// TIA Portal project "Praca_Dyplomowa" (V17)

(* hardware
DEVICE "S7-1200 station_1"  S7-1200 Station
   slot 0: "Rack_0"  S7-1200 Rack  Rack  V1.0
   slot 1: "PLC_1"  CPU 1214C DC/DC/DC  6ES7 214-1AE30-0XB0  V2.2
   slot 3: "AQ 1x12BIT_1"  AQ1 signal board  6ES7 232-4HA30-0XB0  V1.0
DEVICE "HMI_2"  KTP600 Basic color PN
   slot 0: "HMI_2"  KTP600 Basic color PN  6AV6 647-0AD11-3AX0  12.0.0.0
   slot 1: "HMI_RT_2"  KTP600 Basic color PN  6AV6 647-0AD11-3AX0  12.0.0.0
   slot 5: "HMI_2.IE_CP_1"  PROFINET Interface  12.0.0.0
      slot 1: "PROFINET Interface_1"  PROFINET Interface
         slot 1: "Port_1"  Port
*)

// ===== PLC "PLC_1"  CPU 1214C DC/DC/DC =====

VAR_GLOBAL   // PLC tag table "Default tag table"
   "System_Byte" AT %MB1 : Byte;
   "FirstScan" AT %M1.0 : Bool;
   "DiagStatusUpdate" AT %M1.1 : Bool;
   "AlwaysTRUE" AT %M1.2 : Bool;
   "AlwaysFALSE" AT %M1.3 : Bool;
   "Clock_Byte" AT %MB0 : Byte;
   "Clock_10Hz" AT %M0.0 : Bool;
   "Clock_5Hz" AT %M0.1 : Bool;
   "Clock_2.5Hz" AT %M0.2 : Bool;
   "Clock_2Hz" AT %M0.3 : Bool;
   "Clock_1.25Hz" AT %M0.4 : Bool;
   "Clock_1Hz" AT %M0.5 : Bool;
   "Clock_0.625Hz" AT %M0.6 : Bool;
   "Clock_0.5Hz" AT %M0.7 : Bool;
END_VAR

DATA_BLOCK "Dane_Temperatura"   // DB1
{ S7_Optimized_Access := 'FALSE' }
VERSION : 0.1
   VAR
      DS1_DEC : Real;
      DS2_DEC : Real;
      DS3_DEC : Real;
      DS1_DECx100 : Int;
      DS2_DECx100 : Int;
      DS3_DECx100 : Int;
      Przelicznik : Real := 100.0;
      MaxDS_1 : Real;
      MinDS_1 : Real;
      MaxDS_2 : Real := 0.0;
      MinDS_2 : Real := 0.0;
      MaxDS_3 : Real := 0.0;
      MinDS_3 : Real := 0.0;
      MaxDS_1x100 : Int;
      MinDS_1x100 : Int;
      MaxDS_2x100 : Int;
      MinDS_2x100 : Int;
      MaxDS_3x100 : Int;
      MinDS_3x100 : Int;
   END_VAR
BEGIN
END_DATA_BLOCK

DATA_BLOCK "Dane Czujnik Odleglosci"   // DB2
{ S7_Optimized_Access := 'TRUE' }
VERSION : 0.1
   VAR
      Odległość : Int;
   END_VAR
BEGIN
END_DATA_BLOCK

DATA_BLOCK "MB_TCP_Data_Drugi_Serwer"   // DB4
{ S7_Optimized_Access := 'FALSE' }
VERSION : 0.1
   VAR
      IP_serwer_nr_2 : Struct
         Pierwszy_oktet : USInt := 192;
         Drugi_oktet_1 : USInt := 168;
         Trzeci_oktet_2 : USInt := 00;
         Czwarty_oktet_3 : USInt := 251;
      END_STRUCT;
      Port_Serwera_Drugiego : Word := 502;
      Serwer_Drugi : Word := 2;
      Numer_Rejestru : Word := 40001;
      Tryb_Pracy : USInt := 0;
      ILE_danych : Word := 20;
      Data_next_device : Array[1..20] of Word;
      disconnect : Bool;
      przelicznik_cisnienie : Real := 10.0;
      przelicznik_temp : Real := 100.0;
      Cisnieniex10 : Int;
      Tempx100 : Int;
      Cisnienie : Real;
      Temperatura : Real;
      Kod_Błedu : Word;
   END_VAR
BEGIN
END_DATA_BLOCK

DATA_BLOCK "MB_TCP_Data_Trzeci_Serwer"   // DB7
{ S7_Optimized_Access := 'FALSE' }
VERSION : 0.1
   VAR
      IP_serwer_nr_3 : Struct
         Pierwszy_oktet : USInt := 192;
         Drugi_oktet_1 : USInt := 168;
         Trzeci_oktet_2 : USInt := 00;
         Czwarty_oktet_3 : USInt := 252;
      END_STRUCT;
      Port_Serwera_Trzeciego : Word := 502;
      Serwer_Trzeci : Word := 3;
      Numer_Rejestru : Word := 40001;
      Tryb_Pracy : USInt := 0;
      ILE_danych : Word := 20;
      Dane_Trzeci_Serwer : Array[1..20] of Word;
      DISCONNECT : Bool;
      Kod_Błedu : Word;
      Przelicznik_100 : Real := 100.0;
      Przelicznik_1000 : Real := 1000.0;
      ax_1000 : Int;
      ay_1000 : Int;
      az_1000 : Int;
      ax : Real;
      ay : Real;
      az : Real;
      gx_100 : Int;
      gy_100 : Int;
      gz_100 : Int;
      gx : Real;
      gz : Real;
      gy : Real;
      temp_100 : Int;
      temp : Real;
   END_VAR
BEGIN
END_DATA_BLOCK

DATA_BLOCK "MB_SERWER_PLC_DANE"   // DB9
{ S7_Optimized_Access := 'FALSE' }
VERSION : 0.1
   VAR
      DISCONNECT : Bool;
      PLC_serwer_pierwszy : UInt := 5;
      IP_PORT : UInt := 502;
      New_Data_Ready : Bool;
      Data_Read : Bool;
      ERROR : Bool;
      KOD_BLEDU_SERWERA_PLC : Word;
   END_VAR
BEGIN
END_DATA_BLOCK

DATA_BLOCK "MB_TCP_Connection"   // DB10
{ S7_Optimized_Access := 'FALSE' }
VERSION : 0.1
   VAR
      MB_TCP_DISCONNECT : Bool;
      MB_TCP_ERROR : Bool;
      MB_TCP_STATUS : Word;
      MB_TCP_BUSY : Bool;
      MB_TCP_DONE : Bool;
      Connection_Lost : Bool;
   END_VAR
BEGIN
END_DATA_BLOCK

DATA_BLOCK "MB_TCP_Data"   // DB11
{ S7_Optimized_Access := 'FALSE' }
VERSION : 0.1
   VAR
      IP_serwer_nr_1 : Struct
         Pierwszy_oktet : USInt := 192;
         Drugi_oktet_1 : USInt := 168;
         Trzeci_oktet_2 : USInt := 00;
         Czwarty_oktet_3 : USInt := 253;
      END_STRUCT;
      Port_Serwera_Pierwszego : Word := 502;
      Serwer_Pierwszy : Word := 1;
      Numer_Rejestru : Word := 40001;
      Tryb_Pracy : USInt := 0;
      ILE_danych : Word := 26;
      Dane_serwer_pierwszy : Array[1..26] of Word;
   END_VAR
BEGIN
END_DATA_BLOCK

DATA_BLOCK "Zmienne_cyclic_interrupt"   // DB12
{ S7_Optimized_Access := 'TRUE' }
VERSION : 0.1
   VAR RETAIN
      IN : Bool;
      PIN : Bool;
      OUT : Bool;
      POUT : Bool;
      Czas : Time := T#250ms;
   END_VAR
BEGIN
END_DATA_BLOCK

FUNCTION "VL53L1" : Void   // FC1, LAD
{ S7_Optimized_Access := 'TRUE' }
VERSION : 0.1
BEGIN

REGION Network 1
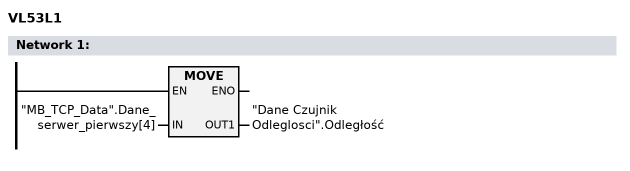
   RUNG wire#powerrail
      { S7_GenerateENO := "TRUE" } Move(in := "MB_TCP_Data".Dane_serwer_pierwszy[4], out1 => "Dane Czujnik Odleglosci".Odległość)
   END_RUNG
   // the same network as SCL:
   "Dane Czujnik Odleglosci".Odległość := "MB_TCP_Data".Dane_serwer_pierwszy[4];
END_REGION
END_FUNCTION

FUNCTION "STATUS_INFO" : Void   // FC2, SCL
{ S7_Optimized_Access := 'TRUE' }
VERSION : 0.1
   VAR_TEMP
      i : Int;
      "a" : Int;
      "b" : Int;
   END_VAR
BEGIN
   IF WORD_TO_INT("MB_TCP_Connection".MB_TCP_STATUS) <> 0 THEN
       "MB_TCP_Connection".Connection_Lost := TRUE;
       FOR #i := 1 TO WORD_TO_INT("MB_TCP_Data".ILE_danych) DO
           "MB_TCP_Data".Dane_serwer_pierwszy[#i] := 0;
       END_FOR;
   ELSE
       "MB_TCP_Connection".Connection_Lost := FALSE;
   END_IF;

   IF WORD_TO_INT("MB_TCP_Data_Drugi_Serwer".Kod_Błedu) <> 0 THEN

       FOR #a := 1 TO WORD_TO_INT("MB_TCP_Data_Trzeci_Serwer".ILE_danych) DO
           "MB_TCP_Data_Drugi_Serwer".Data_next_device[#a] := 0;
       END_FOR;

   END_IF;


   IF WORD_TO_INT("MB_TCP_Data_Trzeci_Serwer".Kod_Błedu) <> 0 THEN

       FOR #b := 1 TO WORD_TO_INT("MB_TCP_Data_Trzeci_Serwer".ILE_danych) DO
           "MB_TCP_Data_Trzeci_Serwer".Dane_Trzeci_Serwer[#b] := 0;
       END_FOR;

   END_IF;
END_FUNCTION

FUNCTION "BMP280" : Void   // FC3, LAD
{ S7_Optimized_Access := 'TRUE' }
VERSION : 0.1
BEGIN

REGION Network 1
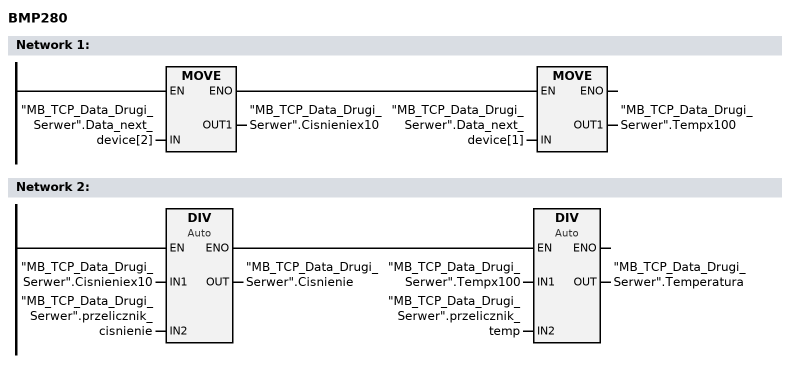
   RUNG wire#powerrail
      { S7_GenerateENO := "TRUE" } Move(in := "MB_TCP_Data_Drugi_Serwer".Data_next_device[2], out1 => "MB_TCP_Data_Drugi_Serwer".Cisnieniex10)
      { S7_GenerateENO := "TRUE" } Move(in := "MB_TCP_Data_Drugi_Serwer".Data_next_device[1], out1 => "MB_TCP_Data_Drugi_Serwer".Tempx100)
   END_RUNG
   // the same network as SCL:
   // ENO of a box is taken as its EN; it also drops when the box reports an error
   "MB_TCP_Data_Drugi_Serwer".Cisnieniex10 := "MB_TCP_Data_Drugi_Serwer".Data_next_device[2];
   "MB_TCP_Data_Drugi_Serwer".Tempx100 := "MB_TCP_Data_Drugi_Serwer".Data_next_device[1];
END_REGION

REGION Network 2
   RUNG wire#powerrail
      { S7_GenerateENO := "TRUE" } Div(in1 := "MB_TCP_Data_Drugi_Serwer".Cisnieniex10, in2 := "MB_TCP_Data_Drugi_Serwer".przelicznik_cisnienie, out => "MB_TCP_Data_Drugi_Serwer".Cisnienie)
      { S7_GenerateENO := "TRUE" } Div(in1 := "MB_TCP_Data_Drugi_Serwer".Tempx100, in2 := "MB_TCP_Data_Drugi_Serwer".przelicznik_temp, out => "MB_TCP_Data_Drugi_Serwer".Temperatura)
   END_RUNG
   // the same network as SCL:
   // ENO of a box is taken as its EN; it also drops when the box reports an error
   "MB_TCP_Data_Drugi_Serwer".Cisnienie := "MB_TCP_Data_Drugi_Serwer".Cisnieniex10 / "MB_TCP_Data_Drugi_Serwer".przelicznik_cisnienie;
   "MB_TCP_Data_Drugi_Serwer".Temperatura := "MB_TCP_Data_Drugi_Serwer".Tempx100 / "MB_TCP_Data_Drugi_Serwer".przelicznik_temp;
END_REGION
END_FUNCTION

FUNCTION "GY521" : Void   // FC4, LAD
{ S7_Optimized_Access := 'TRUE' }
VERSION : 0.1
BEGIN

REGION Network 1
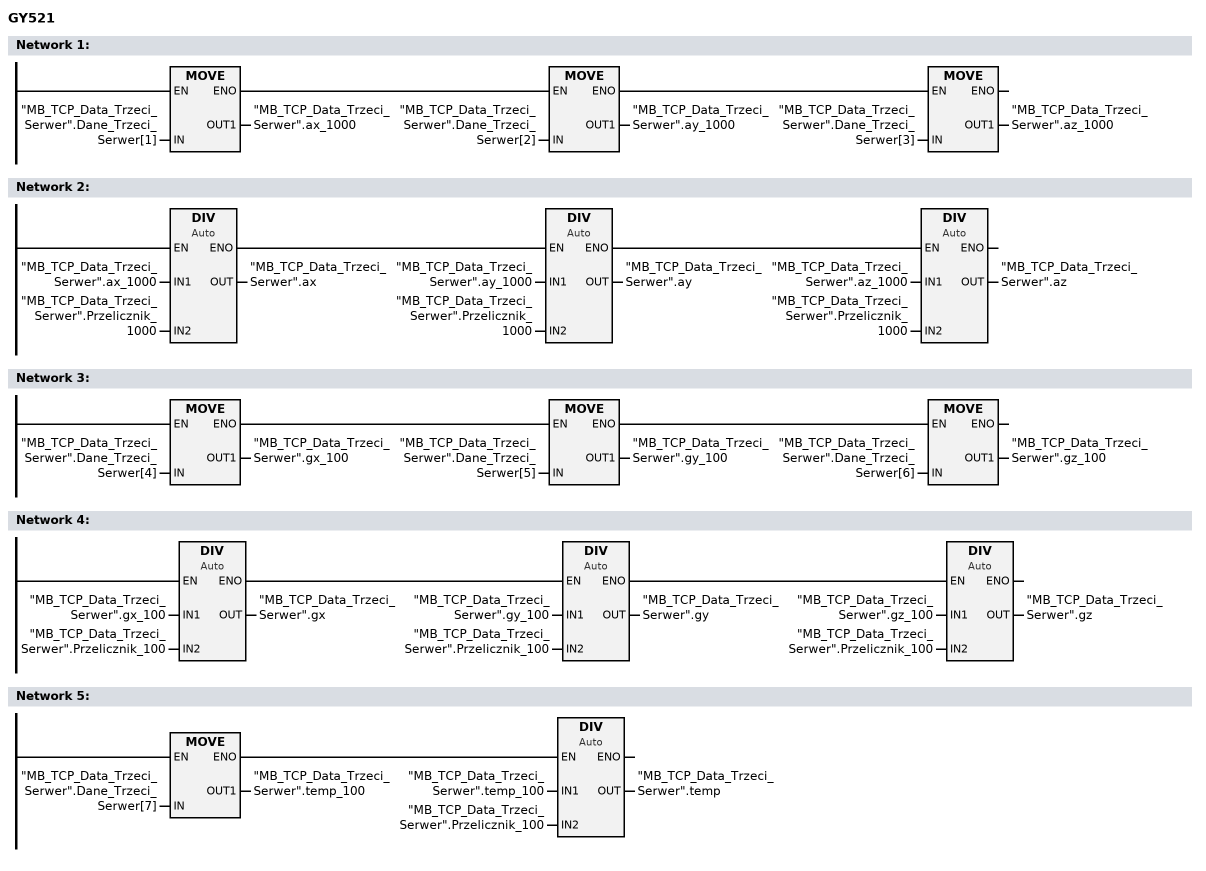
   RUNG wire#powerrail
      { S7_GenerateENO := "TRUE" } Move(in := "MB_TCP_Data_Trzeci_Serwer".Dane_Trzeci_Serwer[1], out1 => "MB_TCP_Data_Trzeci_Serwer".ax_1000)
      { S7_GenerateENO := "TRUE" } Move(in := "MB_TCP_Data_Trzeci_Serwer".Dane_Trzeci_Serwer[2], out1 => "MB_TCP_Data_Trzeci_Serwer".ay_1000)
      { S7_GenerateENO := "TRUE" } Move(in := "MB_TCP_Data_Trzeci_Serwer".Dane_Trzeci_Serwer[3], out1 => "MB_TCP_Data_Trzeci_Serwer".az_1000)
   END_RUNG
   // the same network as SCL:
   // ENO of a box is taken as its EN; it also drops when the box reports an error
   "MB_TCP_Data_Trzeci_Serwer".ax_1000 := "MB_TCP_Data_Trzeci_Serwer".Dane_Trzeci_Serwer[1];
   "MB_TCP_Data_Trzeci_Serwer".ay_1000 := "MB_TCP_Data_Trzeci_Serwer".Dane_Trzeci_Serwer[2];
   "MB_TCP_Data_Trzeci_Serwer".az_1000 := "MB_TCP_Data_Trzeci_Serwer".Dane_Trzeci_Serwer[3];
END_REGION

REGION Network 2
   RUNG wire#powerrail
      { S7_GenerateENO := "TRUE" } Div(in1 := "MB_TCP_Data_Trzeci_Serwer".ax_1000, in2 := "MB_TCP_Data_Trzeci_Serwer".Przelicznik_1000, out => "MB_TCP_Data_Trzeci_Serwer".ax)
      { S7_GenerateENO := "TRUE" } Div(in1 := "MB_TCP_Data_Trzeci_Serwer".ay_1000, in2 := "MB_TCP_Data_Trzeci_Serwer".Przelicznik_1000, out => "MB_TCP_Data_Trzeci_Serwer".ay)
      { S7_GenerateENO := "TRUE" } Div(in1 := "MB_TCP_Data_Trzeci_Serwer".az_1000, in2 := "MB_TCP_Data_Trzeci_Serwer".Przelicznik_1000, out => "MB_TCP_Data_Trzeci_Serwer".az)
   END_RUNG
   // the same network as SCL:
   // ENO of a box is taken as its EN; it also drops when the box reports an error
   "MB_TCP_Data_Trzeci_Serwer".ax := "MB_TCP_Data_Trzeci_Serwer".ax_1000 / "MB_TCP_Data_Trzeci_Serwer".Przelicznik_1000;
   "MB_TCP_Data_Trzeci_Serwer".ay := "MB_TCP_Data_Trzeci_Serwer".ay_1000 / "MB_TCP_Data_Trzeci_Serwer".Przelicznik_1000;
   "MB_TCP_Data_Trzeci_Serwer".az := "MB_TCP_Data_Trzeci_Serwer".az_1000 / "MB_TCP_Data_Trzeci_Serwer".Przelicznik_1000;
END_REGION

REGION Network 3
   RUNG wire#powerrail
      { S7_GenerateENO := "TRUE" } Move(in := "MB_TCP_Data_Trzeci_Serwer".Dane_Trzeci_Serwer[4], out1 => "MB_TCP_Data_Trzeci_Serwer".gx_100)
      { S7_GenerateENO := "TRUE" } Move(in := "MB_TCP_Data_Trzeci_Serwer".Dane_Trzeci_Serwer[5], out1 => "MB_TCP_Data_Trzeci_Serwer".gy_100)
      { S7_GenerateENO := "TRUE" } Move(in := "MB_TCP_Data_Trzeci_Serwer".Dane_Trzeci_Serwer[6], out1 => "MB_TCP_Data_Trzeci_Serwer".gz_100)
   END_RUNG
   // the same network as SCL:
   // ENO of a box is taken as its EN; it also drops when the box reports an error
   "MB_TCP_Data_Trzeci_Serwer".gx_100 := "MB_TCP_Data_Trzeci_Serwer".Dane_Trzeci_Serwer[4];
   "MB_TCP_Data_Trzeci_Serwer".gy_100 := "MB_TCP_Data_Trzeci_Serwer".Dane_Trzeci_Serwer[5];
   "MB_TCP_Data_Trzeci_Serwer".gz_100 := "MB_TCP_Data_Trzeci_Serwer".Dane_Trzeci_Serwer[6];
END_REGION

REGION Network 4
   RUNG wire#powerrail
      { S7_GenerateENO := "TRUE" } Div(in1 := "MB_TCP_Data_Trzeci_Serwer".gx_100, in2 := "MB_TCP_Data_Trzeci_Serwer".Przelicznik_100, out => "MB_TCP_Data_Trzeci_Serwer".gx)
      { S7_GenerateENO := "TRUE" } Div(in1 := "MB_TCP_Data_Trzeci_Serwer".gy_100, in2 := "MB_TCP_Data_Trzeci_Serwer".Przelicznik_100, out => "MB_TCP_Data_Trzeci_Serwer".gy)
      { S7_GenerateENO := "TRUE" } Div(in1 := "MB_TCP_Data_Trzeci_Serwer".gz_100, in2 := "MB_TCP_Data_Trzeci_Serwer".Przelicznik_100, out => "MB_TCP_Data_Trzeci_Serwer".gz)
   END_RUNG
   // the same network as SCL:
   // ENO of a box is taken as its EN; it also drops when the box reports an error
   "MB_TCP_Data_Trzeci_Serwer".gx := "MB_TCP_Data_Trzeci_Serwer".gx_100 / "MB_TCP_Data_Trzeci_Serwer".Przelicznik_100;
   "MB_TCP_Data_Trzeci_Serwer".gy := "MB_TCP_Data_Trzeci_Serwer".gy_100 / "MB_TCP_Data_Trzeci_Serwer".Przelicznik_100;
   "MB_TCP_Data_Trzeci_Serwer".gz := "MB_TCP_Data_Trzeci_Serwer".gz_100 / "MB_TCP_Data_Trzeci_Serwer".Przelicznik_100;
END_REGION

REGION Network 5
   RUNG wire#powerrail
      { S7_GenerateENO := "TRUE" } Move(in := "MB_TCP_Data_Trzeci_Serwer".Dane_Trzeci_Serwer[7], out1 => "MB_TCP_Data_Trzeci_Serwer".temp_100)
      { S7_GenerateENO := "TRUE" } Div(in1 := "MB_TCP_Data_Trzeci_Serwer".temp_100, in2 := "MB_TCP_Data_Trzeci_Serwer".Przelicznik_100, out => "MB_TCP_Data_Trzeci_Serwer".temp)
   END_RUNG
   // the same network as SCL:
   // ENO of a box is taken as its EN; it also drops when the box reports an error
   "MB_TCP_Data_Trzeci_Serwer".temp_100 := "MB_TCP_Data_Trzeci_Serwer".Dane_Trzeci_Serwer[7];
   "MB_TCP_Data_Trzeci_Serwer".temp := "MB_TCP_Data_Trzeci_Serwer".temp_100 / "MB_TCP_Data_Trzeci_Serwer".Przelicznik_100;
END_REGION
END_FUNCTION

FUNCTION "MB_Serwer_PLC" : Void   // FC5, LAD
{ S7_Optimized_Access := 'FALSE' }
VERSION : 0.1
BEGIN

REGION Network 1
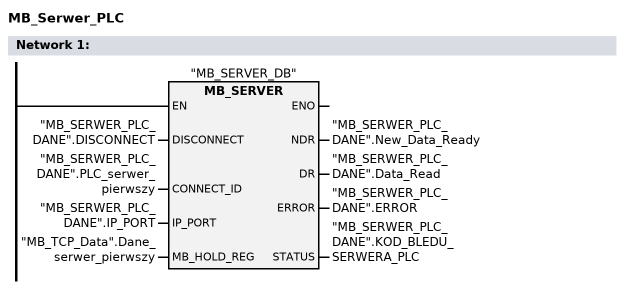
   "MB_SERVER_DB"(DISCONNECT := "MB_SERWER_PLC_DANE".DISCONNECT,   // MB_SERVER
                  CONNECT_ID := "MB_SERWER_PLC_DANE".PLC_serwer_pierwszy,
                  IP_PORT := "MB_SERWER_PLC_DANE".IP_PORT,
                  MB_HOLD_REG := "MB_TCP_Data".Dane_serwer_pierwszy,
                  NDR => "MB_SERWER_PLC_DANE".New_Data_Ready,
                  DR => "MB_SERWER_PLC_DANE".Data_Read,
                  ERROR => "MB_SERWER_PLC_DANE".ERROR,
                  STATUS => "MB_SERWER_PLC_DANE".KOD_BLEDU_SERWERA_PLC);
END_REGION
END_FUNCTION

FUNCTION "FC_BMTCP_Client" : Void   // FC10, LAD
{ S7_Optimized_Access := 'FALSE' }
VERSION : 0.1
BEGIN

REGION Network 1
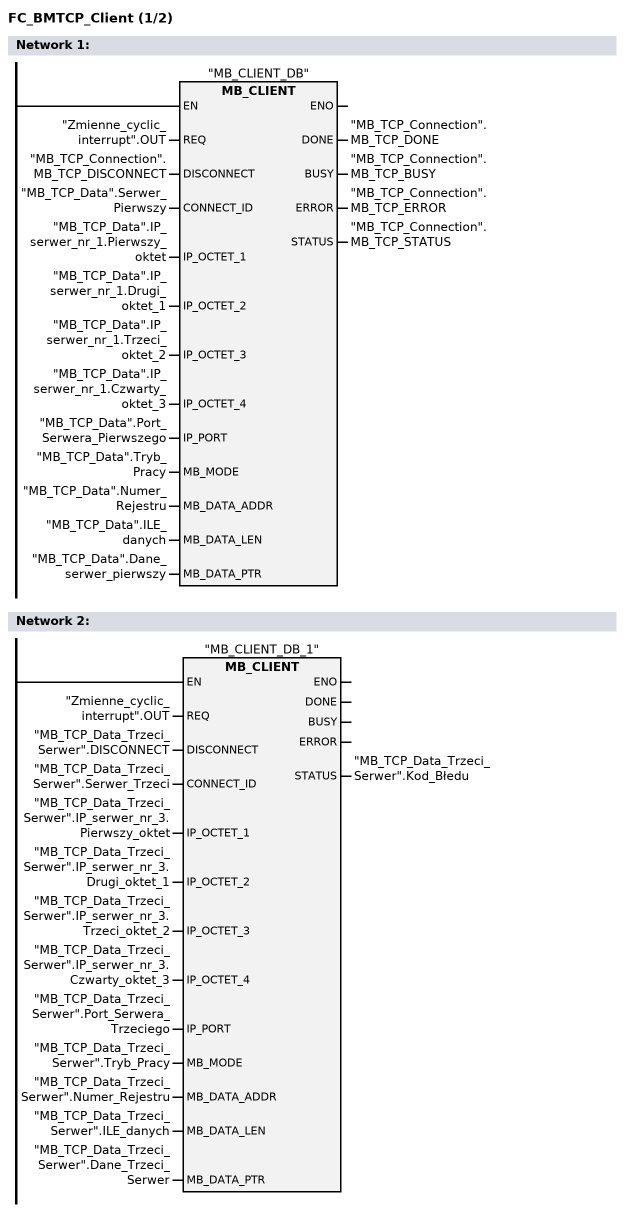
   "MB_CLIENT_DB"(REQ := "Zmienne_cyclic_interrupt".OUT,   // MB_CLIENT
                  DISCONNECT := "MB_TCP_Connection".MB_TCP_DISCONNECT,
                  CONNECT_ID := "MB_TCP_Data".Serwer_Pierwszy,
                  IP_OCTET_1 := "MB_TCP_Data".IP_serwer_nr_1.Pierwszy_oktet,
                  IP_OCTET_2 := "MB_TCP_Data".IP_serwer_nr_1.Drugi_oktet_1,
                  IP_OCTET_3 := "MB_TCP_Data".IP_serwer_nr_1.Trzeci_oktet_2,
                  IP_OCTET_4 := "MB_TCP_Data".IP_serwer_nr_1.Czwarty_oktet_3,
                  IP_PORT := "MB_TCP_Data".Port_Serwera_Pierwszego,
                  MB_MODE := "MB_TCP_Data".Tryb_Pracy,
                  MB_DATA_ADDR := "MB_TCP_Data".Numer_Rejestru,
                  MB_DATA_LEN := "MB_TCP_Data".ILE_danych,
                  MB_DATA_PTR := "MB_TCP_Data".Dane_serwer_pierwszy,
                  DONE => "MB_TCP_Connection".MB_TCP_DONE,
                  BUSY => "MB_TCP_Connection".MB_TCP_BUSY,
                  ERROR => "MB_TCP_Connection".MB_TCP_ERROR,
                  STATUS => "MB_TCP_Connection".MB_TCP_STATUS);
END_REGION

REGION Network 2
   "MB_CLIENT_DB_1"(REQ := "Zmienne_cyclic_interrupt".OUT,   // MB_CLIENT
                    DISCONNECT := "MB_TCP_Data_Trzeci_Serwer".DISCONNECT,
                    CONNECT_ID := "MB_TCP_Data_Trzeci_Serwer".Serwer_Trzeci,
                    IP_OCTET_1 := "MB_TCP_Data_Trzeci_Serwer".IP_serwer_nr_3.Pierwszy_oktet,
                    IP_OCTET_2 := "MB_TCP_Data_Trzeci_Serwer".IP_serwer_nr_3.Drugi_oktet_1,
                    IP_OCTET_3 := "MB_TCP_Data_Trzeci_Serwer".IP_serwer_nr_3.Trzeci_oktet_2,
                    IP_OCTET_4 := "MB_TCP_Data_Trzeci_Serwer".IP_serwer_nr_3.Czwarty_oktet_3,
                    IP_PORT := "MB_TCP_Data_Trzeci_Serwer".Port_Serwera_Trzeciego,
                    MB_MODE := "MB_TCP_Data_Trzeci_Serwer".Tryb_Pracy,
                    MB_DATA_ADDR := "MB_TCP_Data_Trzeci_Serwer".Numer_Rejestru,
                    MB_DATA_LEN := "MB_TCP_Data_Trzeci_Serwer".ILE_danych,
                    MB_DATA_PTR := "MB_TCP_Data_Trzeci_Serwer".Dane_Trzeci_Serwer,
                    STATUS => "MB_TCP_Data_Trzeci_Serwer".Kod_Błedu);
END_REGION

REGION Network 3
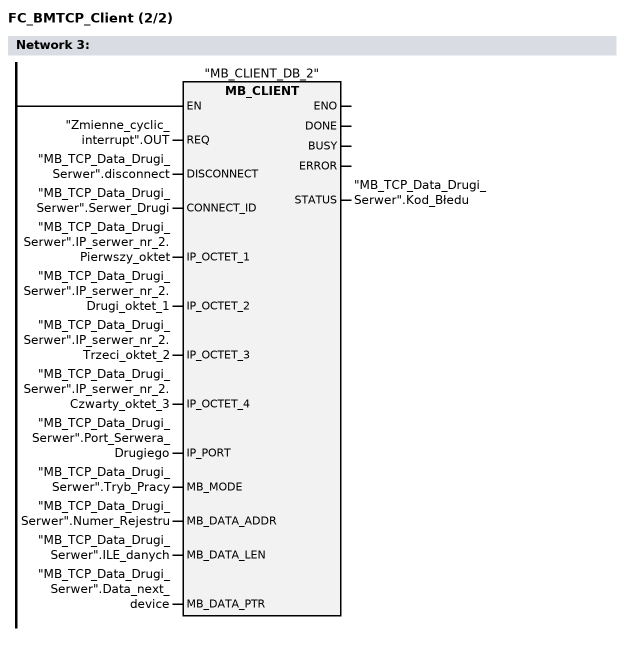
   "MB_CLIENT_DB_2"(REQ := "Zmienne_cyclic_interrupt".OUT,   // MB_CLIENT
                    DISCONNECT := "MB_TCP_Data_Drugi_Serwer".disconnect,
                    CONNECT_ID := "MB_TCP_Data_Drugi_Serwer".Serwer_Drugi,
                    IP_OCTET_1 := "MB_TCP_Data_Drugi_Serwer".IP_serwer_nr_2.Pierwszy_oktet,
                    IP_OCTET_2 := "MB_TCP_Data_Drugi_Serwer".IP_serwer_nr_2.Drugi_oktet_1,
                    IP_OCTET_3 := "MB_TCP_Data_Drugi_Serwer".IP_serwer_nr_2.Trzeci_oktet_2,
                    IP_OCTET_4 := "MB_TCP_Data_Drugi_Serwer".IP_serwer_nr_2.Czwarty_oktet_3,
                    IP_PORT := "MB_TCP_Data_Drugi_Serwer".Port_Serwera_Drugiego,
                    MB_MODE := "MB_TCP_Data_Drugi_Serwer".Tryb_Pracy,
                    MB_DATA_ADDR := "MB_TCP_Data_Drugi_Serwer".Numer_Rejestru,
                    MB_DATA_LEN := "MB_TCP_Data_Drugi_Serwer".ILE_danych,
                    MB_DATA_PTR := "MB_TCP_Data_Drugi_Serwer".Data_next_device,
                    STATUS => "MB_TCP_Data_Drugi_Serwer".Kod_Błedu);
END_REGION
END_FUNCTION

FUNCTION "TEMP_HEX_AND_REAL" : Void   // FC11, LAD
{ S7_Optimized_Access := 'FALSE' }
VERSION : 0.1
BEGIN

REGION Network 1
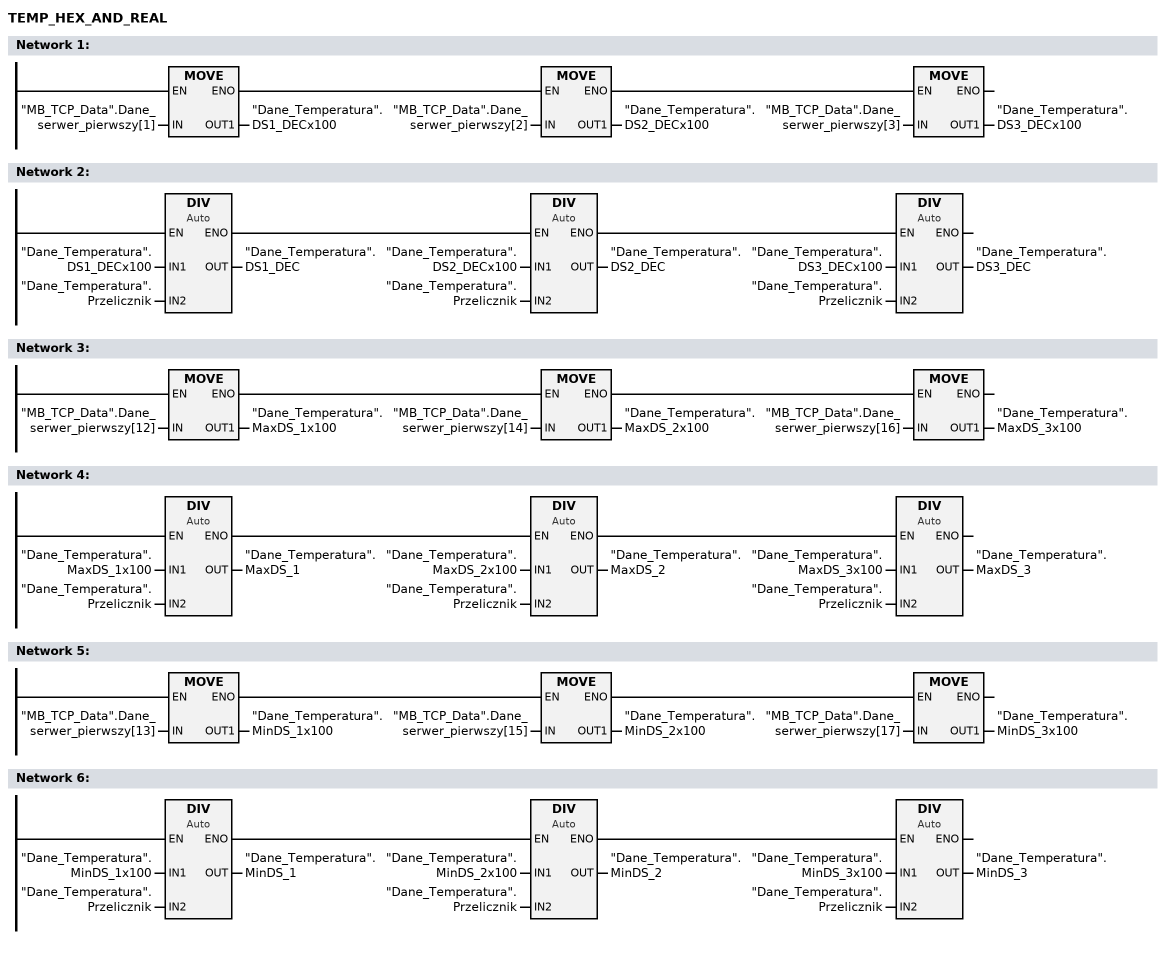
   RUNG wire#powerrail
      { S7_GenerateENO := "TRUE" } Move(in := "MB_TCP_Data".Dane_serwer_pierwszy[1], out1 => "Dane_Temperatura".DS1_DECx100)
      { S7_GenerateENO := "TRUE" } Move(in := "MB_TCP_Data".Dane_serwer_pierwszy[2], out1 => "Dane_Temperatura".DS2_DECx100)
      { S7_GenerateENO := "TRUE" } Move(in := "MB_TCP_Data".Dane_serwer_pierwszy[3], out1 => "Dane_Temperatura".DS3_DECx100)
   END_RUNG
   // the same network as SCL:
   // ENO of a box is taken as its EN; it also drops when the box reports an error
   "Dane_Temperatura".DS1_DECx100 := "MB_TCP_Data".Dane_serwer_pierwszy[1];
   "Dane_Temperatura".DS2_DECx100 := "MB_TCP_Data".Dane_serwer_pierwszy[2];
   "Dane_Temperatura".DS3_DECx100 := "MB_TCP_Data".Dane_serwer_pierwszy[3];
END_REGION

REGION Network 2
   RUNG wire#powerrail
      { S7_GenerateENO := "TRUE" } Div(in1 := "Dane_Temperatura".DS1_DECx100, in2 := "Dane_Temperatura".Przelicznik, out => "Dane_Temperatura".DS1_DEC)
      { S7_GenerateENO := "TRUE" } Div(in1 := "Dane_Temperatura".DS2_DECx100, in2 := "Dane_Temperatura".Przelicznik, out => "Dane_Temperatura".DS2_DEC)
      { S7_GenerateENO := "TRUE" } Div(in1 := "Dane_Temperatura".DS3_DECx100, in2 := "Dane_Temperatura".Przelicznik, out => "Dane_Temperatura".DS3_DEC)
   END_RUNG
   // the same network as SCL:
   // ENO of a box is taken as its EN; it also drops when the box reports an error
   "Dane_Temperatura".DS1_DEC := "Dane_Temperatura".DS1_DECx100 / "Dane_Temperatura".Przelicznik;
   "Dane_Temperatura".DS2_DEC := "Dane_Temperatura".DS2_DECx100 / "Dane_Temperatura".Przelicznik;
   "Dane_Temperatura".DS3_DEC := "Dane_Temperatura".DS3_DECx100 / "Dane_Temperatura".Przelicznik;
END_REGION

REGION Network 3
   RUNG wire#powerrail
      { S7_GenerateENO := "TRUE" } Move(in := "MB_TCP_Data".Dane_serwer_pierwszy[12], out1 => "Dane_Temperatura".MaxDS_1x100)
      { S7_GenerateENO := "TRUE" } Move(in := "MB_TCP_Data".Dane_serwer_pierwszy[14], out1 => "Dane_Temperatura".MaxDS_2x100)
      { S7_GenerateENO := "TRUE" } Move(in := "MB_TCP_Data".Dane_serwer_pierwszy[16], out1 => "Dane_Temperatura".MaxDS_3x100)
   END_RUNG
   // the same network as SCL:
   // ENO of a box is taken as its EN; it also drops when the box reports an error
   "Dane_Temperatura".MaxDS_1x100 := "MB_TCP_Data".Dane_serwer_pierwszy[12];
   "Dane_Temperatura".MaxDS_2x100 := "MB_TCP_Data".Dane_serwer_pierwszy[14];
   "Dane_Temperatura".MaxDS_3x100 := "MB_TCP_Data".Dane_serwer_pierwszy[16];
END_REGION

REGION Network 4
   RUNG wire#powerrail
      { S7_GenerateENO := "TRUE" } Div(in1 := "Dane_Temperatura".MaxDS_1x100, in2 := "Dane_Temperatura".Przelicznik, out => "Dane_Temperatura".MaxDS_1)
      { S7_GenerateENO := "TRUE" } Div(in1 := "Dane_Temperatura".MaxDS_2x100, in2 := "Dane_Temperatura".Przelicznik, out => "Dane_Temperatura".MaxDS_2)
      { S7_GenerateENO := "TRUE" } Div(in1 := "Dane_Temperatura".MaxDS_3x100, in2 := "Dane_Temperatura".Przelicznik, out => "Dane_Temperatura".MaxDS_3)
   END_RUNG
   // the same network as SCL:
   // ENO of a box is taken as its EN; it also drops when the box reports an error
   "Dane_Temperatura".MaxDS_1 := "Dane_Temperatura".MaxDS_1x100 / "Dane_Temperatura".Przelicznik;
   "Dane_Temperatura".MaxDS_2 := "Dane_Temperatura".MaxDS_2x100 / "Dane_Temperatura".Przelicznik;
   "Dane_Temperatura".MaxDS_3 := "Dane_Temperatura".MaxDS_3x100 / "Dane_Temperatura".Przelicznik;
END_REGION

REGION Network 5
   RUNG wire#powerrail
      { S7_GenerateENO := "TRUE" } Move(in := "MB_TCP_Data".Dane_serwer_pierwszy[13], out1 => "Dane_Temperatura".MinDS_1x100)
      { S7_GenerateENO := "TRUE" } Move(in := "MB_TCP_Data".Dane_serwer_pierwszy[15], out1 => "Dane_Temperatura".MinDS_2x100)
      { S7_GenerateENO := "TRUE" } Move(in := "MB_TCP_Data".Dane_serwer_pierwszy[17], out1 => "Dane_Temperatura".MinDS_3x100)
   END_RUNG
   // the same network as SCL:
   // ENO of a box is taken as its EN; it also drops when the box reports an error
   "Dane_Temperatura".MinDS_1x100 := "MB_TCP_Data".Dane_serwer_pierwszy[13];
   "Dane_Temperatura".MinDS_2x100 := "MB_TCP_Data".Dane_serwer_pierwszy[15];
   "Dane_Temperatura".MinDS_3x100 := "MB_TCP_Data".Dane_serwer_pierwszy[17];
END_REGION

REGION Network 6
   RUNG wire#powerrail
      { S7_GenerateENO := "TRUE" } Div(in1 := "Dane_Temperatura".MinDS_1x100, in2 := "Dane_Temperatura".Przelicznik, out => "Dane_Temperatura".MinDS_1)
      { S7_GenerateENO := "TRUE" } Div(in1 := "Dane_Temperatura".MinDS_2x100, in2 := "Dane_Temperatura".Przelicznik, out => "Dane_Temperatura".MinDS_2)
      { S7_GenerateENO := "TRUE" } Div(in1 := "Dane_Temperatura".MinDS_3x100, in2 := "Dane_Temperatura".Przelicznik, out => "Dane_Temperatura".MinDS_3)
   END_RUNG
   // the same network as SCL:
   // ENO of a box is taken as its EN; it also drops when the box reports an error
   "Dane_Temperatura".MinDS_1 := "Dane_Temperatura".MinDS_1x100 / "Dane_Temperatura".Przelicznik;
   "Dane_Temperatura".MinDS_2 := "Dane_Temperatura".MinDS_2x100 / "Dane_Temperatura".Przelicznik;
   "Dane_Temperatura".MinDS_3 := "Dane_Temperatura".MinDS_3x100 / "Dane_Temperatura".Przelicznik;
END_REGION
END_FUNCTION

ORGANIZATION_BLOCK "Main"   // OB1, LAD, ProgramCycle
TITLE = "Main Program Sweep (Cycle)"
{ S7_Optimized_Access := 'TRUE' }
VERSION : 0.1
   VAR_TEMP   // added for the SCL form of the ladder/FBD networks
      _w1 : Bool;
      _w2 : Bool;
      _w3 : Bool;
      _w4 : Bool;
      _w5 : Bool;
   END_VAR
BEGIN

REGION Network 1
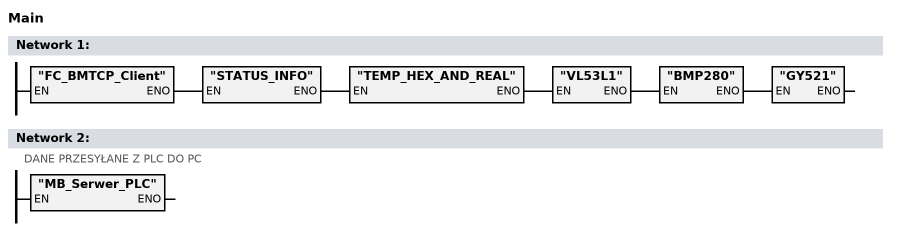
   RUNG wire#powerrail
      "FC_BMTCP_Client"()
      "STATUS_INFO"()
      "TEMP_HEX_AND_REAL"()
      "VL53L1"()
      "BMP280"()
      "GY521"()
   END_RUNG
   // the same network as SCL:
   "FC_BMTCP_Client"(ENO => #_w1);
   "STATUS_INFO"(EN := #_w1, ENO => #_w2);
   "TEMP_HEX_AND_REAL"(EN := #_w2, ENO => #_w3);
   "VL53L1"(EN := #_w3, ENO => #_w4);
   "BMP280"(EN := #_w4, ENO => #_w5);
   IF #_w5 THEN "GY521"(); END_IF;
END_REGION

REGION Network 2
   // DANE PRZESYŁANE Z PLC DO PC
   RUNG wire#powerrail
      "MB_Serwer_PLC"()
   END_RUNG
   // the same network as SCL:
   "MB_Serwer_PLC"();
END_REGION
END_ORGANIZATION_BLOCK

ORGANIZATION_BLOCK "Cyclic interrupt"   // OB30, SCL, CyclicInterrupt
{ S7_Optimized_Access := 'TRUE' }
VERSION : 0.1
BEGIN
   "Zmienne_cyclic_interrupt".OUT := NOT "Zmienne_cyclic_interrupt".OUT;
END_ORGANIZATION_BLOCK

(* ===== HMI "HMI_RT_2" =====
system functions are stored by id; their names below are inferred from use
connection "HMI_Connection_2": ETHERNET, SMART_S7_1200_OMS

HMI tags "Default tag table"
   "Dane_Temperatura_DS1_DEC" : Real = PLC Dane_Temperatura.DS1_DEC AT %DB1.DBD0, 100 ms
   "Dane_Temperatura_DS2_DEC" : Real = PLC Dane_Temperatura.DS2_DEC AT %DB1.DBD4, 100 ms
   "Dane_Temperatura_DS3_DEC" : Real = PLC Dane_Temperatura.DS3_DEC AT %DB1.DBD8, 100 ms
   "Dane Czujnik Odleglosci_Odległość" : Int = PLC "Dane Czujnik Odleglosci".Odległość, 100 ms
   "MB_TCP_Connection_MB_TCP_ERROR" : Bool = PLC MB_TCP_Connection.MB_TCP_ERROR AT %DB10.DBX0.1, 100 ms
   "MB_TCP_Connection_MB_TCP_STATUS" : Word = PLC MB_TCP_Connection.MB_TCP_STATUS AT %DB10.DBW2, 100 ms
   "MB_TCP_Connection_MB_TCP_BUSY" : Bool = PLC MB_TCP_Connection.MB_TCP_BUSY AT %DB10.DBX4.0, 100 ms
   "MB_TCP_Connection_MB_TCP_DONE" : Bool = PLC MB_TCP_Connection.MB_TCP_DONE AT %DB10.DBX4.1, 100 ms
   "MB_TCP_Connection_Connection_Lost" : Bool = PLC MB_TCP_Connection.Connection_Lost AT %DB10.DBX4.2, 100 ms
   "Dane_Temperatura_DS1_DECx100" : Int = PLC Dane_Temperatura.DS1_DECx100 AT %DB1.DBW12, 100 ms
   "Dane_Temperatura_DS2_DECx100" : Int = PLC Dane_Temperatura.DS2_DECx100 AT %DB1.DBW14, 100 ms
   "Dane_Temperatura_DS3_DECx100" : Int = PLC Dane_Temperatura.DS3_DECx100 AT %DB1.DBW16, 100 ms
   "MB_TCP_Data_Static_1[11]" : Word = PLC MB_TCP_Data.Dane_serwer_pierwszy[11] AT %DB11.DBW34, 100 ms
   "MB_TCP_Data_Static_1[10]" : Word = PLC MB_TCP_Data.Dane_serwer_pierwszy[10] AT %DB11.DBW32, 100 ms
   "MB_TCP_Data_Static_1[9]" : Word = PLC MB_TCP_Data.Dane_serwer_pierwszy[9] AT %DB11.DBW30, 100 ms
   "MB_TCP_Data_Static_1[5]" : Word = PLC MB_TCP_Data.Dane_serwer_pierwszy[5] AT %DB11.DBW22, 100 ms
   "MB_TCP_Data_Static_1[6]" : Word = PLC MB_TCP_Data.Dane_serwer_pierwszy[6] AT %DB11.DBW24, 100 ms
   "MB_TCP_Data_Static_1[7]" : Word = PLC MB_TCP_Data.Dane_serwer_pierwszy[7] AT %DB11.DBW26, 100 ms
   "Dane_Temperatura_MaxDS_1" : Real = PLC Dane_Temperatura.MaxDS_1 AT %DB1.DBD22, 100 ms
   "Dane_Temperatura_MaxDS_2" : Real = PLC Dane_Temperatura.MaxDS_2 AT %DB1.DBD30, 100 ms
   "Dane_Temperatura_MaxDS_3" : Real = PLC Dane_Temperatura.MaxDS_3 AT %DB1.DBD38, 100 ms
   "Dane_Temperatura_MinDS_1" : Real = PLC Dane_Temperatura.MinDS_1 AT %DB1.DBD26, 100 ms
   "Dane_Temperatura_MinDS_2" : Real = PLC Dane_Temperatura.MinDS_2 AT %DB1.DBD34, 100 ms
   "Dane_Temperatura_MinDS_3" : Real = PLC Dane_Temperatura.MinDS_3 AT %DB1.DBD42, 100 ms
   "MB_TCP_Data_Static_1[18]" : Word = PLC MB_TCP_Data.Dane_serwer_pierwszy[18] AT %DB11.DBW48, 100 ms
   "MB_TCP_Data_Static_1[21]" : Word = PLC MB_TCP_Data.Dane_serwer_pierwszy[21] AT %DB11.DBW54, 100 ms
   "MB_TCP_Data_Static_1[22]" : Word = PLC MB_TCP_Data.Dane_serwer_pierwszy[22] AT %DB11.DBW56, 100 ms
   "MB_TCP_Data_Static_1[20]" : Word = PLC MB_TCP_Data.Dane_serwer_pierwszy[20] AT %DB11.DBW52, 100 ms
   "MB_TCP_Data_Static_1[19]" : Word = PLC MB_TCP_Data.Dane_serwer_pierwszy[19] AT %DB11.DBW50, 100 ms
   "MB_TCP_Data_next_device_Temperatura" : Real = PLC MB_TCP_Data_Drugi_Serwer.Temperatura AT %DB4.DBD72, 1 s
   "MB_TCP_Data_next_device_Cisnienie" : Real = PLC MB_TCP_Data_Drugi_Serwer.Cisnienie AT %DB4.DBD68, 1 s
   "MB_TCP_Data_Static_1[24]" : Word = PLC MB_TCP_Data.Dane_serwer_pierwszy[24] AT %DB11.DBW60, 100 ms
   "MB_TCP_Data_Static_1[25]" : Word = PLC MB_TCP_Data.Dane_serwer_pierwszy[25] AT %DB11.DBW62, 100 ms
   "MB_TCP_Data_Static_1[23]" : Word = PLC MB_TCP_Data.Dane_serwer_pierwszy[23] AT %DB11.DBW58, 100 ms
   "MB_TCP_Data_Dane_serwer_pierwszy[26]" : Word = PLC MB_TCP_Data.Dane_serwer_pierwszy[26] AT %DB11.DBW64, 1 s
   "MB_TCP_Data_Drugi_Serwer_Kod_Błedu" : Word = PLC MB_TCP_Data_Drugi_Serwer.Kod_Błedu AT %DB4.DBW76, 1 s
   "MB_TCP_Data_Trzeci_Serwer_temp" : Real = PLC MB_TCP_Data_Trzeci_Serwer.temp AT %DB7.DBD104, 100 ms
   "MB_TCP_Data_Trzeci_Serwer_gx" : Real = PLC MB_TCP_Data_Trzeci_Serwer.gx AT %DB7.DBD90, 100 ms
   "MB_TCP_Data_Trzeci_Serwer_ax" : Real = PLC MB_TCP_Data_Trzeci_Serwer.ax AT %DB7.DBD72, 100 ms
   "MB_TCP_Data_Trzeci_Serwer_az" : Real = PLC MB_TCP_Data_Trzeci_Serwer.az AT %DB7.DBD80, 100 ms
   "MB_TCP_Data_Trzeci_Serwer_ay" : Real = PLC MB_TCP_Data_Trzeci_Serwer.ay AT %DB7.DBD76, 100 ms
   "MB_TCP_Data_Trzeci_Serwer_gy" : Real = PLC MB_TCP_Data_Trzeci_Serwer.gy AT %DB7.DBD98, 100 ms
   "MB_TCP_Data_Trzeci_Serwer_gz" : Real = PLC MB_TCP_Data_Trzeci_Serwer.gz AT %DB7.DBD94, 100 ms
   "MB_TCP_Data_Trzeci_Serwer_Kod_Błedu" : Word = PLC MB_TCP_Data_Trzeci_Serwer.Kod_Błedu AT %DB7.DBW56, 100 ms

screen "Screen_1" 320x240
   TextField "Text field_1" at 78,11 size 39x16; Text 'TEMP.'
   IOField "I/O field_3" at 72,78 size 70x23; FormatPattern s999.99
      ProcessValue <- "Dane_Temperatura_DS3_DEC"
   TextField "Text field_2" at 20,11 size 52x16; Text 'CZUJNIK'
   TextField "Text field_3" at 33,32 size 31x16; Text 'Nr. 1'
   TextField "Text field_4" at 33,56 size 31x16; Text 'Nr. 2'
   TextField "Text field_5" at 33,78 size 31x16; Text 'Nr. 3'
   IOField "I/O field_1" at 72,54 size 70x23; FormatPattern s999.99
      ProcessValue <- "Dane_Temperatura_DS2_DEC"
   IOField "I/O field_2" at 72,30 size 70x23; FormatPattern s999.99
      ProcessValue <- "Dane_Temperatura_DS1_DEC"
   TextField "Text field_6" at 124,32 size 16x16; Text '°C'
   TextField "Text field_7" at 124,56 size 16x16; Text '°C'
   TextField "Text field_8" at 123,80 size 16x16; Text '°C'
   TextField "Text field_9" at 8,138 size 114x16; Text 'Odczyt Odległości:'
   IOField "I/O field_4" at 232,137 size 62x23; FormatPattern 9999
      ProcessValue <- "Dane Czujnik Odleglosci_Odległość"
   TextField "Text field_10" at 274,141 size 20x13; Text 'mm'
   TextField "Text field_11" at 186,11 size 115x16; Text 'STAN POŁĄCZENIA'
   TextField "Text field_12" at 185,33 size 46x15; Text 'STATUS'
   TextField "Text field_13" at 185,51 size 58x15; Text 'Kod Błędu'
   TextField "Text field_14" at 186,72 size 92x15; Text 'Trwa zapytanie'
   GraphicView "Graphic view_1" at 231,34 size 17x16; Picture "Graphic_1"
      Visibility <- "MB_TCP_Connection_Connection_Lost"
   GraphicView "Graphic view_2" at 230,33 size 18x16; Picture "Graphic_2"
      Visibility <- "MB_TCP_Connection_Connection_Lost"
   IOField "I/O field_5" at 251,51 size 58x17; FormatPattern FFFF
      ProcessValue <- "MB_TCP_Connection_MB_TCP_STATUS"
   TextField "Text field_16" at 185,84 size 73x15; Text 'Modbus TCP'
   Circle "Circle_1" at 286,75 size 24x24
      Appearance <- "MB_TCP_Connection_MB_TCP_BUSY"
   TextField "Text field_15" at 7,114 size 216x16; Text 'Liczba wykrytych czujników temp :'
   IOField "I/O field_6" at 232,113 size 62x23; FormatPattern 99999
      ProcessValue <- "MB_TCP_Data_Static_1[18]"
   TextField "Text field_17" at 7,165 size 166x16; Text 'Odczyt Natężenia Dźwięku:'
   IOField "I/O field_7" at 232,163 size 63x23; FormatPattern 99999
      ProcessValue <- "MB_TCP_Data_Static_1[23]"
   Button "Button_1" at 8,196 size 96x32; TextOff 'DC18B20 Nr 1'
      on Click: ActivateScreen("Przebieg_DC1", 0)
   Button "Button_2" at 113,196 size 96x32; TextOff 'DC18B20 Nr 2'
      on Activate: ActivateScreen("Przebieg_DC2", 0)
   Button "Button_3" at 217,196 size 96x32; TextOff 'DC18B20 Nr 3'
      on Activate: ActivateScreen("Przebieg_DC3", 0)

screen "Screen_2" 320x240
   TextField "Text field_1" at 66,0 size 66x15; Text 'T. Aktualna'
   IOField "I/O field_3" at 153,19 size 70x23; FormatPattern s999999999.99
      ProcessValue <- "Dane_Temperatura_MaxDS_1"
   TextField "Text field_2" at 6,2 size 43x15; Text 'Czujnik'
   TextField "Text field_3" at 15,23 size 31x16; Text 'Nr. 1'
   IOField "I/O field_2" at 68,19 size 70x23; FormatPattern s999999999.99
      ProcessValue <- "Dane_Temperatura_DS1_DEC"
   TextField "Text field_6" at 121,22 size 16x16; Text '°C'
   TextField "Text field_11" at 161,0 size 48x15; Text 'T. Maks.'
   TextField "Text field_12" at 248,0 size 38x15; Text 'T. Min.'
   TextField "Text field_13" at 9,46 size 74x15; Text 'Alarm Temp.'
   TextField "Text field_14" at 121,47 size 90x15; Text 'Status Czujnika'
   Circle "Circle_1" at 85,47 size 24x24
      Appearance <- "MB_TCP_Data_Static_1[5]"
   TextField "Text field_4" at 11,59 size 57x12; Text '-10°C || 80°C'
   Circle "Circle_2" at 221,47 size 24x24
      Appearance <- "MB_TCP_Data_Static_1[9]"
   TextField "Text field_7" at 205,23 size 16x16; Text '°C'
   IOField "I/O field_1" at 240,19 size 70x23; FormatPattern s999999999.99
      ProcessValue <- "Dane_Temperatura_MinDS_1"
   TextField "Text field_8" at 293,23 size 16x16; Text '°C'
   TextField "Text field_5" at 66,77 size 66x15; Text 'T. Aktualna'
   IOField "I/O field_4" at 153,96 size 70x23; FormatPattern s999999999.99
      ProcessValue <- "Dane_Temperatura_MaxDS_2"
   TextField "Text field_9" at 6,79 size 43x15; Text 'Czujnik'
   TextField "Text field_10" at 15,100 size 31x16; Text 'Nr. 2'
   IOField "I/O field_5" at 68,96 size 70x23; FormatPattern s999999999.99
      ProcessValue <- "Dane_Temperatura_DS2_DEC"
   TextField "Text field_15" at 121,99 size 16x16; Text '°C'
   TextField "Text field_16" at 161,77 size 48x15; Text 'T. Maks.'
   TextField "Text field_17" at 248,77 size 38x15; Text 'T. Min.'
   TextField "Text field_18" at 9,123 size 74x15; Text 'Alarm Temp.'
   TextField "Text field_19" at 121,124 size 90x15; Text 'Status Czujnika'
   Circle "Circle_3" at 85,124 size 24x24
      Appearance <- "MB_TCP_Data_Static_1[6]"
   TextField "Text field_20" at 11,136 size 57x12; Text '-10°C || 80°C'
   Circle "Circle_4" at 221,124 size 24x24
      Appearance <- "MB_TCP_Data_Static_1[10]"
   TextField "Text field_21" at 205,100 size 16x16; Text '°C'
   IOField "I/O field_6" at 240,96 size 70x23; FormatPattern s999999999.99
      ProcessValue <- "Dane_Temperatura_MinDS_2"
   TextField "Text field_22" at 293,100 size 16x16; Text '°C'
   TextField "Text field_23" at 66,160 size 66x15; Text 'T. Aktualna'
   IOField "I/O field_7" at 153,179 size 70x23; FormatPattern s999999999.99
      ProcessValue <- "Dane_Temperatura_MaxDS_3"
   TextField "Text field_24" at 6,162 size 43x15; Text 'Czujnik'
   TextField "Text field_25" at 15,179 size 31x16; Text 'Nr. 3'
   IOField "I/O field_8" at 68,179 size 70x23; FormatPattern s999999999.99
      ProcessValue <- "Dane_Temperatura_DS3_DEC"
   TextField "Text field_26" at 121,182 size 16x16; Text '°C'
   TextField "Text field_27" at 161,160 size 48x15; Text 'T. Maks.'
   TextField "Text field_28" at 248,160 size 38x15; Text 'T. Min.'
   TextField "Text field_29" at 11,204 size 74x15; Text 'Alarm Temp.'
   TextField "Text field_30" at 125,209 size 90x15; Text 'Status Czujnika'
   Circle "Circle_5" at 90,207 size 24x24
      Appearance <- "MB_TCP_Data_Static_1[7]"
   TextField "Text field_31" at 9,218 size 57x12; Text '-10°C || 80°C'
   Circle "Circle_6" at 221,206 size 24x24
      Appearance <- "MB_TCP_Data_Static_1[11]"
      Visibility <- "MB_TCP_Data_Static_1[11]"
   TextField "Text field_32" at 205,183 size 16x16; Text '°C'
   IOField "I/O field_9" at 240,179 size 70x23; FormatPattern s999999999.99
      ProcessValue <- "Dane_Temperatura_MinDS_3"
   TextField "Text field_33" at 293,183 size 16x16; Text '°C'

screen "Screen_3" 320x240
   TextField "Text field_1" at 78,11 size 10x16; Text 'Text'
   IOField "I/O field_3" at 159,78 size 70x23; FormatPattern 99999
      ProcessValue <- "MB_TCP_Data_Static_1[22]"
   TextField "Text field_2" at 94,5 size 112x16; Text 'Czujnik Odległości'
   TextField "Text field_3" at 31,33 size 69x16; Text 'Odległość :'
   TextField "Text field_4" at 31,56 size 102x16; Text 'Max. Odległość :'
   TextField "Text field_5" at 31,78 size 99x16; Text 'Min. Odległość:'
   IOField "I/O field_1" at 159,56 size 70x23; FormatPattern 99999
      ProcessValue <- "MB_TCP_Data_Static_1[21]"
   IOField "I/O field_2" at 159,33 size 70x23; FormatPattern s9999
      ProcessValue <- "Dane Czujnik Odleglosci_Odległość"
   IOField "I/O field_6" at 157,126 size 72x23; FormatPattern 99999
      ProcessValue <- "MB_TCP_Data_Static_1[20]"
   TextField "Text field_6" at 33,125 size 112x20; Text 'Liczba Detali :'
   TextField "Text field_7" at 34,178 size 106x16; Text 'Status Czujnika:'
   Circle "Circle_1" at 177,172 size 29x29
      Appearance <- "MB_TCP_Data_Static_1[19]"
   TextField "Text field_10" at 205,81 size 20x13; Text 'mm'
   TextField "Text field_8" at 205,59 size 20x13; Text 'mm'
   TextField "Text field_9" at 206,36 size 20x13; Text 'mm'
   TextField "Text field_11" at 209,131 size 16x13; Text 'szt'

screen "Screen_4" 320x240
   TrendView "Trend view_1" at 0,23 size 319x167
   IOField "I/O field_2" at 68,204 size 96x23; FormatPattern 99999
      ProcessValue <- "MB_TCP_Data_Static_1[25]"
   TextField "Text field_2" at 107,2 size 110x16; Text 'Czujnik MAX4466'
   TextField "Text field_28" at 13,199 size 40x15; Text 'Liczba'
   TextField "Text field_30" at 171,205 size 90x15; Text 'Status Czujnika'
   TextField "Text field_1" at 8,212 size 53x15; Text 'Zgłoszeń'
   Circle "Circle_1" at 274,198 size 29x29
      Appearance <- "MB_TCP_Data_Dane_serwer_pierwszy[26]"

screen "Screen_5" 320x240
   IOField "I/O field_3" at 132,80 size 70x23; FormatPattern 99999.9
      ProcessValue <- "MB_TCP_Data_next_device_Cisnienie"
   TextField "Text field_4" at 31,56 size 84x16; Text 'Temperatura:'
   TextField "Text field_5" at 31,78 size 59x16; Text 'Ciśnienie:'
   IOField "I/O field_1" at 133,53 size 70x23; FormatPattern s999.99
      ProcessValue <- "MB_TCP_Data_next_device_Temperatura"
   TextField "Text field_10" at 176,84 size 21x13; Text 'hPa'
   TextField "Text field_2" at 106,3 size 102x16; Text 'Serwer numer II'
   TextField "Text field_7" at 184,54 size 16x16; Text '°C'
   TextField "Text field_13" at 32,108 size 58x15; Text 'Kod Błędu'
   IOField "I/O field_5" at 132,108 size 69x19; FormatPattern FFFF
      ProcessValue <- "MB_TCP_Data_Drugi_Serwer_Kod_Błedu"

screen "Screen_6" 320x240
   TextField "Text field_2" at 106,3 size 107x16; Text 'Serwer numer III'
   TextField "Text field_4" at 13,48 size 84x16; Text 'Temperatura:'
   IOField "I/O field_1" at 107,48 size 77x19; FormatPattern s999.99
      ProcessValue <- "MB_TCP_Data_Trzeci_Serwer_temp"
   TextField "Text field_7" at 160,48 size 16x16; Text '°C'
   TextField "Text field_5" at 20,81 size 62x16; Text 'Żyroskop:'
   TextField "Text field_1" at 13,102 size 17x16; Text 'gx'
   TextField "Text field_3" at 13,125 size 17x16; Text 'gy'
   TextField "Text field_6" at 13,150 size 16x16; Text 'gz'
   TextField "Text field_8" at 166,126 size 16x16; Text 'ay'
   TextField "Text field_9" at 167,100 size 16x16; Text 'ax'
   TextField "Text field_10" at 166,148 size 15x16; Text 'az'
   IOField "I/O field_2" at 41,101 size 77x19; FormatPattern s999.99
      ProcessValue <- "MB_TCP_Data_Trzeci_Serwer_gx"
   IOField "I/O field_3" at 41,126 size 77x19; FormatPattern s999.99
      ProcessValue <- "MB_TCP_Data_Trzeci_Serwer_gy"
   IOField "I/O field_4" at 41,150 size 77x19; FormatPattern s999.99
      ProcessValue <- "MB_TCP_Data_Trzeci_Serwer_gz"
   TextField "Text field_12" at 183,80 size 83x16; Text 'Akcelerometr'
   IOField "I/O field_5" at 195,102 size 77x19; FormatPattern s999.999
      ProcessValue <- "MB_TCP_Data_Trzeci_Serwer_ax"
   IOField "I/O field_6" at 195,125 size 77x19; FormatPattern s999.999
      ProcessValue <- "MB_TCP_Data_Trzeci_Serwer_ay"
   IOField "I/O field_7" at 195,149 size 77x19; FormatPattern s999.999
      ProcessValue <- "MB_TCP_Data_Trzeci_Serwer_az"
   TextField "Text field_13" at 21,192 size 58x15; Text 'Kod Błędu'
   IOField "I/O field_8" at 91,191 size 69x19; FormatPattern FFFF
      ProcessValue <- "MB_TCP_Data_Trzeci_Serwer_Kod_Błedu"
   TextField "Text field_11" at 256,102 size 10x16; Text 'g'
   TextField "Text field_14" at 256,125 size 10x16; Text 'g'
   TextField "Text field_15" at 256,148 size 10x16; Text 'g'
   TextField "Text field_16" at 94,101 size 21x16; Text '°/s'
   TextField "Text field_17" at 95,126 size 21x16; Text '°/s'
   TextField "Text field_18" at 94,149 size 21x16; Text '°/s'

screen "Przebieg_DC1" 320x240
   TrendView "Trend view_1" at 0,23 size 319x167
   TextField "Text field_2" at 86,1 size 136x16; Text 'Czujnik DC18B20 nr 1'
   Button "Button_1" at 207,200 size 96x32; TextOff 'Powrót'
      on Click: function_efd93a16()

screen "Przebieg_DC2" 320x240
   TrendView "Trend view_1" at 0,23 size 319x167
   TextField "Text field_2" at 86,1 size 136x16; Text 'Czujnik DC18B20 nr 2'
   Button "Button_1" at 207,200 size 96x32; TextOff 'Powrót'
      on Click: function_efd93a16()

screen "Przebieg_DC3" 320x240
   TrendView "Trend view_1" at 0,23 size 319x167
   TextField "Text field_2" at 86,1 size 136x16; Text 'Czujnik DC18B20 nr 3'
   Button "Button_1" at 207,200 size 96x32; TextOff 'Powrót'
      on Click: function_efd93a16()
*)